
   Warranty conditions, liability, AND support -
      IF the application has been made available free OF charge, the following applies:
      * We DO NOT provide a warranty FOR Any OF the information contained in this document.
      * All other rights AND claims against Siemens AG irrespective OF legal basis are excluded. In particular claims FOR damages against Siemens AG 
      in the CASE OF Product outage, downtime, loss OF profit, either directly, indirectly OR consequential damage are excluded.
      * This does NOT apply when liability is compulsory BY law, e. g. in the CASE OF the Product liability act, premeditation, an act OF gross negligence 
      BY superiors AND managerial staff OF Siemens AG OR in cases OF fraudulent concealment OF defects.
      * This limitation OF liability also applies TO sub-contractors, suppliers, delegates, superiors AND managerial staff OF Siemens AG.
      German law shall apply TO this agreement FOR customers with head offices in Germany; Swiss law FOR customers with head offices outside Germany. 
      Application OF the United Nations Convention on Contracts FOR the International Sale OF Goods as OF 11.04.1980 (CISG) is excluded.
   *)

   // ===========================================================================
   //  Begin the LOGIC section:

   // Determine the Number of Sts_Events for given alarm/warning area
   // // S7-300 Logic:
   // UDT_Event = 66 bytes in length
   // S7-300 Logic:
   //#tempAnyPointer := #Sts_EventSummation.Sts_Events;    // temp Any Pointer for FC_ArrrayLength call.
   //"FC_ArrayLength"(ArraySource:= #tempAnyPointer, ArrayLength:=66, SIZE=> #Sts_EventSummation.Wrk_EventArraySize);
   // S7-1500 Logic:
   // "FC_ArrayLength_S7-1500"(Array_ToBe_Sized := #Sts_EventSummation.Sts_Events,
      //                      ArraySize => #Sts_EventSummation.Wrk_EventArraySize);

   // Cleanup the summation - This FB is to be called after the numerous "FB_PMLe_EventSum" calls.
   IF #Prev_NumAllEvents > #Sts_EventSummation.Sts_NumEvents THEN
       FOR #Index := #Sts_EventSummation.Sts_NumEvents TO (#Prev_NumAllEvents-1) DO
             #Sts_EventSummation.Sts_Events[#Index]:= #ZeroEvent;   // clear the first out event
       END_FOR;
   END_IF;

   #Prev_NumAllEvents := #Sts_EventSummation.Sts_NumEvents;     

   #Sts_EventSummation.Sts_Category_0_Latched := #Sts_EventSummation.Wrk_Category_0_Latched;
   #Sts_EventSummation.Sts_Category_1_Latched := #Sts_EventSummation.Wrk_Category_1_Latched;
   #Sts_EventSummation.Sts_Category_2_Latched := #Sts_EventSummation.Wrk_Category_2_Latched;
   #Sts_EventSummation.Sts_Category_3_Latched := #Sts_EventSummation.Wrk_Category_3_Latched;
   #Sts_EventSummation.Sts_Category_4_Latched := #Sts_EventSummation.Wrk_Category_4_Latched;
   #Sts_EventSummation.Sts_Category_6_Latched := #Sts_EventSummation.Wrk_Category_5_Latched;
   #Sts_EventSummation.Sts_Category_7_Latched := #Sts_EventSummation.Wrk_Category_6_Latched;
   #Sts_EventSummation.Sts_Category_8_Latched := #Sts_EventSummation.Wrk_Category_8_Latched;
   #Sts_EventSummation.Sts_Category_9_Latched := #Sts_EventSummation.Wrk_Category_9_Latched;

   #Sts_EventSummation.Sts_Category_0_NotLatched := #Sts_EventSummation.Wrk_Category_0_NotLatched;
   #Sts_EventSummation.Sts_Category_1_NotLatched := #Sts_EventSummation.Wrk_Category_1_NotLatched;
   #Sts_EventSummation.Sts_Category_2_NotLatched := #Sts_EventSummation.Wrk_Category_2_NotLatched;
   #Sts_EventSummation.Sts_Category_3_NotLatched := #Sts_EventSummation.Wrk_Category_3_NotLatched;
   #Sts_EventSummation.Sts_Category_4_NotLatched := #Sts_EventSummation.Wrk_Category_4_NotLatched;
   #Sts_EventSummation.Sts_Category_6_NotLatched := #Sts_EventSummation.Wrk_Category_5_NotLatched;
   #Sts_EventSummation.Sts_Category_7_NotLatched := #Sts_EventSummation.Wrk_Category_6_NotLatched;
   #Sts_EventSummation.Sts_Category_8_NotLatched := #Sts_EventSummation.Wrk_Category_8_NotLatched;
   #Sts_EventSummation.Sts_Category_9_NotLatched := #Sts_EventSummation.Wrk_Category_9_NotLatched;

   #Sts_EventSummation.Sts_CurrentActiveEvent  := #Sts_EventSummation.Wrk_CurrentActiveEvent; 

   //  ------------------------------------------------------------------

   ENO:= true;   // Set the ENO output
END_FUNCTION_BLOCK

FUNCTION_BLOCK "FB_TR88_CPG_EventSortFilter"   // FB3106, SCL
TITLE = PackML Event Sort Filter (TR88 CPG Template)
{ S7_Optimized_Access := 'TRUE' }
AUTHOR : FoodBev
FAMILY : ISATR88e
NAME : EvSrtFlt
VERSION : 1.21
// Sorts and filters event data. It can filter and only show events in a certain category, can sort by time, and can group by category
   VAR_INPUT
      Cmd_FilterActiveEvents : Bool;
      Cmd_FilterCategory : Bool;
      Cfg_FilterCategory : Int;
      Cmd_Sort : Bool;
      Cfg_SortCategory : Bool;
   END_VAR
   VAR_OUTPUT
      Sts_SortFilterNumEvents : Int;
   END_VAR
   VAR_IN_OUT
      In_Events : Array[0.."TR88_CPG_NoOfStsElements_EventSum"] of "UDT_TR88_CPG_Event";   // 30 Events - matches UDT declaration
      In_NumEvents : Int;
      Sts_SortFilterEventList : Array[0.."TR88_CPG_NoOfHMISortEvents"] of "UDT_TR88_CPG_Event";   // 20 Filtered Events
   END_VAR
   VAR
      Compare_True : Bool;
      temp_DT_1 : Date_And_Time;   // Temp Date & Time value #1 - Siemens
      temp_DT_2 : Date_And_Time;   // Temp Date & Time value #2 - Siemens
      FilterAcknowledged : Bool;
      FilterActive : Bool;
      FilterCategory : Bool;
      Index : Int;   // was DINT
      Index_End : Int;   // was DINT
      Index_NumEvents : Int;   // was DINT
      Index_Start : Int;   // was DINT
      MaxSize : Int;   // was DINT
      Prev_NumEvents : Int;   // was DINT
      siftDown_Child : Int;   // was DINT
      siftDown_End : Int;   // was DINT
      siftDown_Root : Int;   // was DINT
      TempEvent : "UDT_TR88_CPG_Event";
      ZeroEvent : "UDT_TR88_CPG_Event";
      Index_2 : Int;   // Index value used for DO and FOR loops
      Compare_1 : Bool;   // Siemens. Compare of TimeEvents #1
      Compare_2 : Bool;   // Siemens. Compare of TimeEvents #2
      SortingEventStatus : Array[0..29] of "UDT_TR88_CPG_Event";   // Added for V1.2
      SortingNumEventsStatus : Int;   // Added for V1.2
   END_VAR
   VAR_TEMP
      tempAnyPointer : DInt;
      siftDown_LeftChild : Int;
      siftDown_RightChild : Int;
   END_VAR
BEGIN
   // ============================================================================ 
   // FUNCTION_BLOCK "FB_PMLe_EventSortFilter"    
   // ---------------------------------------------------------------------------
   // Siemens Industry, Inc.
   // Food & Beverage VSS
   // ---------------------------------------------------------------------------
   // FUNCTIONALITY:  
   // Function Block to control Event Sort Filter commands
   // ---------------------------------------------------------------------------
   // change log table:
   // version        date          expert in charge        changes applied
   // 
   //  1.2         2012-08-20          M.Pieper             Matches Rev 1.2
   //  1.21       2015-01-27           M.Pieper            Updated S7-1500 Array Size Logic.
   // ===========================================================================
   (*
   THIS SOFTWARE IS PROVIDED "AS IS" AND WITHOUT WARRANTIES OF ANY KIND, WHETHER EXPRESS OR IMPLIED.

   General information -
       Note :  the standard applications are NOT binding AND DO NOT claim TO be complete regarding configuration, equipment OR any eventuality which may arise. 
       The standard applications DO NOT represent specific customer solutions, but are only intended TO provide support FOR typical tasks. You are responsible 
       FOR the proper operation OF the described products. These standard applications DO NOT relieve you OF your responsibility regarding the safe handling 
       when using, installing operating AND maintaining the equipment. BY using these standard applications, you agree that Siemens cannot be made liable FOR 
       possible damage beyond the mentioned liability clause. We reserve the right TO make changes AND revisions TO these standard applications at Any Time 
       without prior notice. In the CASE OF Any differences between the suggestions made in these standard applications AND other publications from Siemens, 
       such as catalogs, the contents OF the other documentation have priority.

   Warranty conditions, liability, AND support -
      IF the application has been made available free OF charge, the following applies:
      * We DO NOT provide a warranty FOR Any OF the information contained in this document.
      * All other rights AND claims against Siemens AG irrespective OF legal basis are excluded. In particular claims FOR damages against Siemens AG 
      in the CASE OF Product outage, downtime, loss OF profit, either directly, indirectly OR consequential damage are excluded.
      * This does NOT apply when liability is compulsory BY law, e. g. in the CASE OF the Product liability act, premeditation, an act OF gross negligence 
      BY superiors AND managerial staff OF Siemens AG OR in cases OF fraudulent concealment OF defects.
      * This limitation OF liability also applies TO sub-contractors, suppliers, delegates, superiors AND managerial staff OF Siemens AG.
      German law shall apply TO this agreement FOR customers with head offices in Germany; Swiss law FOR customers with head offices outside Germany. 
      Application OF the United Nations Convention on Contracts FOR the International Sale OF Goods as OF 11.04.1980 (CISG) is excluded.
   *)

   // ===========================================================================
   //  Begin the LOGIC section:
   // Event Sort and Filter
   // Determine the Number of Events for given alarm/warning area
   // UDT_Event = 66 bytes in length 
   // S7-300 Code:
   // #tempAnyPointer := #Sts_SortFilterEventList;    // temp Any Pointer for FC_ArrrayLength call.
   // "FC_ArrayLength"(ArraySource :=  #tempAnyPointer, ArrayLength := 66, SIZE =>  #MaxSize);
   // S7-1500 Code:
   "FC_ArrayLength_S7-1500"(Array_ToBe_Sized := #Sts_SortFilterEventList,
                            ArraySize => #MaxSize);

   IF #In_NumEvents < #MaxSize - 1 THEN
       #SortingNumEventsStatus := DINT_TO_INT(#In_NumEvents);
   ELSE
       #SortingNumEventsStatus := #MaxSize - 1;
   END_IF;

   // Filter
   IF #Cmd_FilterCategory OR #Cmd_FilterActiveEvents THEN
       #Index_NumEvents := 0;
       FOR #Index := 0 TO (#SortingNumEventsStatus - 1) DO         // Siemens added DINT_TO_INT   // should be "In_NumEvents-1"
           #FilterCategory := FALSE;
           #FilterAcknowledged := FALSE;
           #FilterActive := FALSE;
           IF #Cmd_FilterCategory AND (#In_Events[#Index].Category = #Cfg_FilterCategory) THEN
               #FilterCategory := 1;
           END_IF;

           IF #Cmd_FilterActiveEvents AND (#In_Events[#Index].Trigger) THEN
               #FilterActive := 1;
           END_IF;

           IF ((#Cmd_FilterCategory AND #FilterCategory) OR NOT (#Cmd_FilterCategory)) AND ((#Cmd_FilterActiveEvents AND #FilterActive) OR NOT (#Cmd_FilterActiveEvents)) THEN
               #SortingEventStatus[#Index_NumEvents] := #In_Events[#Index];
               #Index_NumEvents := #Index_NumEvents + 1;
           END_IF;

           IF (#Index_NumEvents >= #SortingNumEventsStatus) THEN
               EXIT;
           END_IF;
       END_FOR;

       #SortingNumEventsStatus := #Index_NumEvents;

       // ELSE COP(In_Events[0],Sts_SortFilterEventList[0],Sts_SortFilterNumEvents
   ELSE
       FOR #Index_2 := 0 TO #SortingNumEventsStatus - 1 DO
           #SortingEventStatus[#Index_2] := #In_Events[#Index_2];
       END_FOR;                                            // End FOR loop
   END_IF;                                                 // End Cmd_FilterCategory OR Cmd_FilterActiveEvents THEN....


   // Heap Sort #1
   IF #Cmd_Sort THEN
       // Initial Heapify
       #Index_Start := (#SortingNumEventsStatus / 2);         //-1;
       WHILE #Index_Start >= 0 DO
           // siftDown logic
           #siftDown_Root := #Index_Start;
           #siftDown_End := #SortingNumEventsStatus - 1;
           #siftDown_LeftChild := #siftDown_Root * 2 + 1;
           #siftDown_RightChild := #siftDown_Root * 2 + 2;
           WHILE (#siftDown_LeftChild) <= #siftDown_End DO //while left child exists, find which child is greatest
               IF (#siftDown_LeftChild) = #siftDown_End THEN  // if this is the last element, use it
                   #siftDown_Child := #siftDown_LeftChild;
               ELSIF #Cfg_SortCategory AND (#SortingEventStatus[#siftDown_LeftChild].Category > #SortingEventStatus[#siftDown_RightChild].Category) THEN
                   // if sorting by category, use highest category
                   #siftDown_Child := #siftDown_LeftChild;
               ELSIF (#Cfg_SortCategory AND (#SortingEventStatus[#siftDown_LeftChild].Category = #SortingEventStatus[#siftDown_RightChild].Category)) OR NOT (#Cfg_SortCategory) THEN
                   // if both children are the same cat or no sorting by cat, sort by date
                   #temp_DT_1 := #SortingEventStatus[#siftDown_LeftChild].DateTime;   // Date & Time of Event.TimeEvent[Heap]
                   #temp_DT_2 := #SortingEventStatus[#siftDown_RightChild].DateTime; // Date & Time of Event.TimeEvent[Heap+1]          
                   IF #temp_DT_1 > #temp_DT_2 THEN                                      // is [siftDown_Root*2].TimeEvent > [siftDown_Root*2+1].TimeEvent
                       #siftDown_Child := #siftDown_LeftChild;
                   ELSE
                       #siftDown_Child := #siftDown_RightChild;
                   END_IF;  // END_IF "DT1 > DT2
               ELSE
                   #siftDown_Child := #siftDown_RightChild; // this happens if right.cat > left.cat and sorting by cat
               END_IF; // END_IF "(siftDown_Root*2)..."

               //compare if root and child need to be swapped
               //swap if root has lower category or earlier date
               #Compare_True := 0;
               IF #Cfg_SortCategory AND (#SortingEventStatus[#siftDown_Root].Category < #SortingEventStatus[#siftDown_Child].Category) THEN
                   #Compare_True := 1;
               ELSIF (#Cfg_SortCategory AND (#SortingEventStatus[#siftDown_Root].Category = #SortingEventStatus[#siftDown_Child].Category))
                   OR NOT (#Cfg_SortCategory) THEN
                   #temp_DT_1 := #SortingEventStatus[#siftDown_Root].DateTime;   // Date & Time of Event.TimeEvent[Heap]
                   #temp_DT_2 := #SortingEventStatus[#siftDown_Child].DateTime;  // Date & Time of Event.TimeEvent[Heap+1] 
                   IF #temp_DT_1 < #temp_DT_2 THEN                                  // is [siftDown_Root].TimeEvent < [siftDown_Root+1].TimeEvent
                       #Compare_True := 1;
                   END_IF;  // END_IF "IF Compare_1 ..."           
               END_IF; //END_IF "IF Cfg_SortCategory AND (.."

               IF #Compare_True THEN
                   #TempEvent := #SortingEventStatus[#siftDown_Root];
                   #SortingEventStatus[#siftDown_Root] := #SortingEventStatus[#siftDown_Child];
                   #SortingEventStatus[#siftDown_Child] := #TempEvent;
                   #siftDown_Root := #siftDown_Child;
                   #siftDown_LeftChild := #siftDown_Root * 2 + 1;
                   #siftDown_RightChild := #siftDown_Root * 2 + 2;
               ELSE
                   EXIT;
               END_IF;

           END_WHILE;
           #Index_Start := #Index_Start - 1;
       END_WHILE;

       // Heap Sort #2
       #Index_End := #SortingNumEventsStatus - 1;
       WHILE #Index_End >= 1 DO
           #TempEvent := #SortingEventStatus[0];
           #SortingEventStatus[0] := #SortingEventStatus[#Index_End];
           #SortingEventStatus[#Index_End] := #TempEvent;
           // siftDown
           #siftDown_Root := 0;
           #siftDown_End := #Index_End - 1;
           #siftDown_LeftChild := #siftDown_Root * 2 + 1;
           #siftDown_RightChild := #siftDown_Root * 2 + 2;
           WHILE (#siftDown_LeftChild) <= #siftDown_End DO
               IF (#siftDown_LeftChild) = #siftDown_End THEN
                   #siftDown_Child := #siftDown_LeftChild;
               ELSIF #Cfg_SortCategory AND (#SortingEventStatus[#siftDown_LeftChild].Category > #SortingEventStatus[#siftDown_RightChild].Category) THEN
                   #siftDown_Child := #siftDown_LeftChild;
               ELSIF (#Cfg_SortCategory AND (#SortingEventStatus[#siftDown_LeftChild].Category = #SortingEventStatus[#siftDown_RightChild].Category)) OR NOT (#Cfg_SortCategory) THEN
                   #temp_DT_1 := #SortingEventStatus[#siftDown_LeftChild].DateTime;
                   #temp_DT_2 := #SortingEventStatus[#siftDown_RightChild].DateTime;

                   IF #temp_DT_1 > #temp_DT_2 THEN
                       #siftDown_Child := #siftDown_LeftChild;
                   ELSE
                       #siftDown_Child := #siftDown_RightChild;
                   END_IF;
               ELSE
                   #siftDown_Child := #siftDown_RightChild;
               END_IF;

               #Compare_True := FALSE;
               IF #Cfg_SortCategory AND (#SortingEventStatus[#siftDown_Root].Category < #SortingEventStatus[#siftDown_Child].Category) THEN
                   #Compare_True := TRUE;
               ELSIF (#Cfg_SortCategory AND (#SortingEventStatus[#siftDown_Root].Category = #SortingEventStatus[#siftDown_Child].Category)) OR NOT (#Cfg_SortCategory) THEN
                   #temp_DT_1 := #SortingEventStatus[#siftDown_Root].DateTime;
                   #temp_DT_2 := #SortingEventStatus[#siftDown_Child].DateTime;

                   IF #temp_DT_1 < #temp_DT_2 THEN
                       #Compare_True := TRUE;
                   END_IF;
               END_IF;

               IF #Compare_True THEN
                   #TempEvent := #SortingEventStatus[#siftDown_Root];
                   #SortingEventStatus[#siftDown_Root] := #SortingEventStatus[#siftDown_Child];
                   #SortingEventStatus[#siftDown_Child] := #TempEvent;
                   #siftDown_Root := #siftDown_Child;
                   #siftDown_LeftChild := #siftDown_Root * 2 + 1;
                   #siftDown_RightChild := #siftDown_Root * 2 + 2;
               ELSE
                   EXIT;
               END_IF;
           END_WHILE;
           #Index_End := #Index_End - 1;
       END_WHILE;
   END_IF; //END_IF -> IF Cmd_Sort THEN"

   // Copy SortingEventStatus (working area) to Sts_SortFilterEventList (out)
   // FOR Index  := 0  TO SortingNumEventsStatus DO   
   FOR #Index := 0 TO #SortingNumEventsStatus - 1 DO
       #Sts_SortFilterEventList[#Index] := #SortingEventStatus[#Index];
   END_FOR;
   // End FOR loop
   #Sts_SortFilterNumEvents := #SortingNumEventsStatus;

   // Clean up event list
   IF #Prev_NumEvents > #Sts_SortFilterNumEvents THEN
       //FOR Index  :=  Sts_SortFilterNumEvents TO Prev_NumEvents-1 DO
       FOR #Index := #Sts_SortFilterNumEvents TO #Prev_NumEvents DO
           #Sts_SortFilterEventList[#Index] := #ZeroEvent;
       END_FOR;
   END_IF;

   #Prev_NumEvents := #Sts_SortFilterNumEvents;

   // End of Main Logic.
   //----------------------------------------------------- 

   ENO := true;   // Set the ENO output
END_FUNCTION_BLOCK

FUNCTION_BLOCK "FB_TR88_CPG_Msg_Scroll"   // FB3108, SCL
TITLE = PackML HMI Message Scroll (TR88 CPG Template)
{ S7_Optimized_Access := 'TRUE' }
AUTHOR : FoodBev
FAMILY : ISATR88e
NAME : MsgScrll
VERSION : 1.0
   VAR_INPUT
      Trigger : Bool;   // input trigger to enable scroll logic
      NumEvents : Int;   // input value with number of active events
      In_Events : Array[0.."TR88_CPG_NoOfHMISortEvents"] of "UDT_TR88_CPG_Event";   // incoming events list
   END_VAR
   VAR_OUTPUT
      Msg_Scroll : String[40];   // message output value
   END_VAR
   VAR
      Scroll_Index : Int;   // index value for scroll logic
      TriggerOS : Bool;
      MaxSize : Int;   // was DINT
   END_VAR
   VAR_TEMP
      Scroll_Index_Max : Int;
   END_VAR
BEGIN
   // ============================================================================ 
   // FUNCTION_BLOCK "FB_PMLe_Msg_Scroll"    
   // ---------------------------------------------------------------------------
   // Siemens Industry, Inc.
   // Food & Beverage VMM
   // ---------------------------------------------------------------------------
   // functionality:
   // Function Block used to scoll messages from an array of EVENT to a single
   // ---------------------------------------------------------------------------
   // change log table:
   // version        date          expert in charge        changes applied
   // 
   // 1.0         2012-02-28          M.Pieper           Matches Rev 1.0
   // 1.01        2015-04-01          M.Pieper          Changed "In_Events" from array size of [0..19]
   //                                                    to Array[0.."CPG_TR88_NoOfHMISortEvents"]
   // ===========================================================================
   (*
   THIS SOFTWARE IS PROVIDED "AS IS" AND WITHOUT WARRANTIES OF ANY KIND, WHETHER EXPRESS OR IMPLIED.

   General information -
       Note :  the standard applications are NOT binding AND DO NOT claim TO be complete regarding configuration, equipment OR any eventuality which may arise. 
       The standard applications DO NOT represent specific customer solutions, but are only intended TO provide support FOR typical tasks. You are responsible 
       FOR the proper operation OF the described products. These standard applications DO NOT relieve you OF your responsibility regarding the safe handling 
       when using, installing operating AND maintaining the equipment. BY using these standard applications, you agree that Siemens cannot be made liable FOR 
       possible damage beyond the mentioned liability clause. We reserve the right TO make changes AND revisions TO these standard applications at Any Time 
       without prior notice. In the CASE OF Any differences between the suggestions made in these standard applications AND other publications from Siemens, 
       such as catalogs, the contents OF the other documentation have priority.

   Warranty conditions, liability, AND support -
      IF the application has been made available free OF charge, the following applies:
      * We DO NOT provide a warranty FOR Any OF the information contained in this document.
      * All other rights AND claims against Siemens AG irrespective OF legal basis are excluded. In particular claims FOR damages against Siemens AG 
      in the CASE OF Product outage, downtime, loss OF profit, either directly, indirectly OR consequential damage are excluded.
      * This does NOT apply when liability is compulsory BY law, e. g. in the CASE OF the Product liability act, premeditation, an act OF gross negligence 
      BY superiors AND managerial staff OF Siemens AG OR in cases OF fraudulent concealment OF defects.
      * This limitation OF liability also applies TO sub-contractors, suppliers, delegates, superiors AND managerial staff OF Siemens AG.
      German law shall apply TO this agreement FOR customers with head offices in Germany; Swiss law FOR customers with head offices outside Germany. 
      Application OF the United Nations Convention on Contracts FOR the International Sale OF Goods as OF 11.04.1980 (CISG) is excluded.
   *)

   // ===========================================================================
   //  Begin the LOGIC section:
   "FC_ArrayLength_S7-1500"(Array_ToBe_Sized := #In_Events,
                            ArraySize => #MaxSize);

   IF #NumEvents > #MaxSize THEN
       #Scroll_Index_Max := #MaxSize;
   ELSE
       #Scroll_Index_Max := #NumEvents;
   END_IF;

   // Statement Section 
   IF #Trigger AND NOT #TriggerOS THEN
       #Scroll_Index := #Scroll_Index + 1;  // increment the indext
       IF  #Scroll_Index > #Scroll_Index_Max - 1 THEN
               #Scroll_Index := 0;
           END_IF;
      #Msg_Scroll := #In_Events[#Scroll_Index].Message;      // move the message from the UDT_Event structure to string output.  

       #TriggerOS := TRUE;              // Set the trigger OS bit
   END_IF;

   IF NOT #Trigger AND #TriggerOS THEN
       #TriggerOS := FALSE;
   END_IF;

   ENO:= true;   // Set the ENO output
END_FUNCTION_BLOCK

FUNCTION_BLOCK "FB_TR88_CPG_OEE"   // FB3109, SCL
TITLE = PackML Real-Time OEE Calculation (TR88 CPG Template)
{ S7_Optimized_Access := 'TRUE' }
AUTHOR : FoodBev
FAMILY : ISATR88
NAME : OEE
VERSION : 1.1
   VAR_INPUT
      TotalProdProcessed : DInt;   // Total Number OF Products Processed
      TotalDefectiveProd : DInt;   // Total Number OF Defective Products
      TimeSinceLastReset : DInt;   // Total Acumulative TIME since Last RESET
      MachineDesignSpeed : Real;   // Machine Design Speed
   END_VAR
   VAR_OUTPUT
      OEE_RealTimeValue : Real;   // REAL TIME OEE value (availabilty x performance x quality)
      OEE_Availability : Real;   // OEE - Availability value
      OEE_Performance : Real;   // OEE - Performance value
      OEE_Quality : Real;   // OEE - Quality value
   END_VAR
   VAR_IN_OUT
      ModeCumulativeTimes : Array[0.."LPMLV30_MODES_UPPER_LIM"] of DInt;   // Mode Cummulative Times
   END_VAR
   VAR
      TotalProdProcessed_In : DInt;   // Initial "TotalProdProcessed" value after accum TIME reset
      TotalDefectiveProd_In : DInt;   // Initial "TotalDefectiveProcessed" value after accum TIME reset
      AcumTimeEqualZero : Bool;   // The "TimeSinceLastReset" is = 0 seconds
      AcumTimeEqualZeroOS : Bool;   // OneShot for "TimeSinceLastReset" is = 0 seconds
   END_VAR
   VAR_TEMP
      temp_TimeSinceLastReset : Real;   // used to eliminate divide by zero errors
      temp_TotalProducts : Real;   // used to eliminate divide by zero errors
      temp_DefectiveProducts : Real;   // used to eliminate divide by zero errors
   END_VAR
BEGIN
   // ============================================================================ 
   // FUNCTION_BLOCK "FB_PML_OEE"    
   // ---------------------------------------------------------------------------
   // Siemens Industry, Inc.
   // Food & Beverage VSS
   // ---------------------------------------------------------------------------
   // functionality: Function Block to calculate real-time OEE values
   // ---------------------------------------------------------------------------
   // change log table:
   // version        date          expert in charge        changes applied
   // 
   //  1.00         2012-02-28          M.Pieper        Original - using OEE Realtime calculation
   //  1.10         2012-09-04          M.Pieper        Added seperate Availabity, Performace, Quality calculation
   //  1.20         2014-07-07          M.Pieper        Updated interface FOR new Mode/State FB          
   //  1.201        2016-03-01          M.Pieper        Added logic to prevent floating point / divide by zero errors
   //  // ===========================================================================
   (*
   THIS SOFTWARE IS PROVIDED "AS IS" AND WITHOUT WARRANTIES OF ANY KIND, WHETHER EXPRESS OR IMPLIED.

   General information -
       Note :  the standard applications are NOT binding AND DO NOT claim TO be complete regarding configuration, equipment OR any eventuality which may arise. 
       The standard applications DO NOT represent specific customer solutions, but are only intended TO provide support FOR typical tasks. You are responsible 
       FOR the proper operation OF the described products. These standard applications DO NOT relieve you OF your responsibility regarding the safe handling 
       when using, installing operating AND maintaining the equipment. BY using these standard applications, you agree that Siemens cannot be made liable FOR 
       possible damage beyond the mentioned liability clause. We reserve the right TO make changes AND revisions TO these standard applications at Any Time 
       without prior notice. In the CASE OF Any differences between the suggestions made in these standard applications AND other publications from Siemens, 
       such as catalogs, the contents OF the other documentation have priority.

   Warranty conditions, liability, AND support -
      IF the application has been made available free OF charge, the following applies:
      * We DO NOT provide a warranty FOR Any OF the information contained in this document.
      * All other rights AND claims against Siemens AG irrespective OF legal basis are excluded. In particular claims FOR damages against Siemens AG 
      in the CASE OF Product outage, downtime, loss OF profit, either directly, indirectly OR consequential damage are excluded.
      * This does NOT apply when liability is compulsory BY law, e. g. in the CASE OF the Product liability act, premeditation, an act OF gross negligence 
      BY superiors AND managerial staff OF Siemens AG OR in cases OF fraudulent concealment OF defects.
      * This limitation OF liability also applies TO sub-contractors, suppliers, delegates, superiors AND managerial staff OF Siemens AG.
      German law shall apply TO this agreement FOR customers with head offices in Germany; Swiss law FOR customers with head offices outside Germany. 
      Application OF the United Nations Convention on Contracts FOR the International Sale OF Goods as OF 11.04.1980 (CISG) is excluded.
   *)

   // ===========================================================================
   //  Begin the LOGIC section:
   //  
   (* ISA TR88.00.02 Document - 9.1 OEE Definition:
   Overall Equipment Effectiveness (OEE) is a measure comparing how well manufacturing equipment is running compared to the ideal plant. The resulting measurement is expressed as the ratio of the actual
   output of the equipment divided by the maximum possible output of the equipment under ideal conditions. OEE is calculated by multiplying three independently measured values: Availability,
   Performance Rate, and Quality Rate. The fundamental OEE definition is defined as an availability ratio multiplied by a performance ratio multiplied by a quality ratio.

   OEE = Availability x Performance x Quality

   Where each component is defined as the following:
   Availability = Operating Time / Planned Production Time
   Performance = Total Pieces / (Operating Time* Ideal Run Rate)
   Quality = Good Pieces / Total Pieces

   OEE is often displayed as a waterfall object in which the major components of Availability, Performance, and Quality are displayed graphically.
   *)

   // Determine is TimeSinceLastReset value is equal to zero.
   IF  #TimeSinceLastReset   = 0 THEN
       #AcumTimeEqualZero   := TRUE;  // SET the AcumTimeEqualZero bool tag
   ELSE
       #AcumTimeEqualZero   := FALSE; // RESET the AcumTimeEqualZero bool tag
       #AcumTimeEqualZeroOS := FALSE; // RESET the AcumTimeEqualZero one-shot bool tag
   END_IF;

   // Update the AcumTimeEqualZeroOS One-Shot bool
   IF #AcumTimeEqualZero AND NOT #AcumTimeEqualZeroOS THEN
      #AcumTimeEqualZeroOS := TRUE;  // Set the One-Shot bool tag
   END_IF;

   // Update the inital product count values after the accum timer value has been reset
   IF #AcumTimeEqualZeroOS THEN
      #TotalProdProcessed_In := #TotalProdProcessed;
      #TotalDefectiveProd_In := #TotalDefectiveProd;
   END_IF;  

   // Update the TimeSinceLastReset temp. value.  If = 0 (zero) then change to 0.0001 to ensure no divide by zero errors
   IF #TimeSinceLastReset = 0 THEN
       #temp_TimeSinceLastReset := 0.0001;
   ELSE
       #temp_TimeSinceLastReset := DINT_TO_REAL(#TimeSinceLastReset);
   END_IF;

   (*  9.1.1 Availability Definition
   Availability is defined as operating time divided by planned production time. The basic concept behind availability is to show the time the machine has been running divided by the time that the
   machine has been planned to run. Typical losses in this area are losses to unplanned maintenance, cleaning, changeovers, and breakdowns.
   * Availability = Operating Time / Planned Production Time Operating Time is defined as the amount of time the machine has been attempting to produce parts.  
   * Planned Production Time is defined as the total amount of time the machine has been scheduled to run. 
   *)
   // Availablity = operating time (attempt to run production) / planned production time
   #OEE_Availability :=   DINT_TO_REAL (#ModeCumulativeTimes[1]) / #temp_TimeSinceLastReset;
   IF #OEE_Availability > 1 THEN #OEE_Availability := 1.0; END_IF;
   IF #OEE_Availability < 0 THEN #OEE_Availability := 0.0; END_IF;

   (* 9.1.2 Performance Definition
   Performance is defined as the total number of pieces on which the machine operated divided by the ideal production if a machine ran perfectly for the allocated amount of operating time.
   * Performance = Total Pieces / (Operating Time* Ideal Run Rate).  
   * Total Pieces is defined as good pieces and bad pieces during the production run. This should be linked to the main consumed count of the machine. If a filler, this should be bottles into the filler.
   * Operating Time is defined as the amount of time the machine has been attempting to produce parts. (Same as above)
   * Ideal Run Rate is defined as the ideal rate that the machine can run for the product that is being run on the machine and the way the machine is configured.
   *)
   // Performance = Total Pieces / (Operating Time * Ideal Run Rate / 60)
   #OEE_Performance := (DINT_TO_REAL(#TotalProdProcessed-#TotalProdProcessed_In))/((#temp_TimeSinceLastReset * #MachineDesignSpeed/60.0));
   IF #OEE_Performance > 1 THEN #OEE_Performance := 1.0; END_IF;
   IF #OEE_Performance < 0 THEN #OEE_Performance := 0.0; END_IF;

   (*  9.1.3 Quality Definition
   Quality is defined as the total number of good pieces divided by the total number of pieces on which the machine operated.
   * Quality = Good Pieces / Total Pieces
   * Good Pieces is defined as only good pieces processed during the production run. So this is the main production processed count of the machine. If a filler, this should be bottles out of the filler.
   * Total Pieces includes good pieces and bad pieces during the production run. This should be linked to the main consumed count of the machine. 
      If a filler, this should be bottles into the filler. This should be the same count as used in the performance definition.
   *)
   // Quality = Good Piece / Total Piece
   #temp_TotalProducts     :=  DINT_TO_REAL(#TotalProdProcessed-#TotalProdProcessed_In);
   #temp_DefectiveProducts :=  DINT_TO_REAL(#TotalDefectiveProd-#TotalDefectiveProd_In);

   // Prevent divide by zero errors by checking if Total Products <> 0.0
   IF (#TotalProdProcessed-#TotalProdProcessed_In) = 0 THEN 
       #temp_TotalProducts := 0.0001;
   END_IF;

   // Make sure that defective products < total products
   IF #temp_DefectiveProducts > #temp_TotalProducts THEN
       #temp_DefectiveProducts := 0.0;
   END_IF;

   #OEE_Quality            := (#temp_TotalProducts - #temp_DefectiveProducts) / #temp_TotalProducts;
   IF #OEE_Quality  > 1 THEN #OEE_Quality  := 1.0; END_IF;
   IF #OEE_Quality  < 0 THEN #OEE_Quality  := 0.0; END_IF;
   IF #temp_TotalProducts  = 0 THEN #OEE_Quality  := 0.0; END_IF;

   // OEE_ReatTimeValue := ((DINT_TO_REAL(TotalProdProcessed-TotalProdProcessed_Initial) - DINT_TO_REAL(TotalDefectiveProd-TotalDefectiveProd_Initial)) / ((DINT_TO_REAL(TimeSinceLastReset) * MachineDesignSpeed/60.0)));
   #OEE_RealTimeValue := #OEE_Availability * #OEE_Performance * #OEE_Quality;

   // End of Main Logic.
   ENO:= true;   // Set the ENO output
END_FUNCTION_BLOCK

FUNCTION_BLOCK "FB_TR88_CPG_AlarmMove"   // FB3110, SCL
TITLE = PackML Alarm Move
{ S7_Optimized_Access := 'TRUE' }
AUTHOR : FoodBev
FAMILY : ISATR88e
NAME : AlrmMov
VERSION : 1.01
// ------------------------------------------------------------------------------------------
//   Begin the variable declartion section ....
//  Block Parameters
   VAR_INPUT
      Sts_NumEvents : Int;   // Number OF Active Alarms
   END_VAR
   VAR_OUTPUT
      Sts_error : Bool;   // Error Status. 0=no error, 1=error
      Sts_errorCode : Int;   // Error code /number
   END_VAR
   VAR_IN_OUT
      Source : Array[0.."TR88_CPG_NoOfStsElements_EventSum"] of "UDT_TR88_CPG_Event";   // source location of the machine alarms
      Destination : Array[0.."TR88_CPG_NoOfPackTagsAdminEvents"] of "UDT_TR88_CPG_Event";   // destination location of the PackTag alarms
   END_VAR
   VAR
      Source_NumEvents : Int;   // MAX # OF Events - source event list
      Destination_NumEvents : Int;   // MAX # OF Events - destination event list
      Index : Int;   // index value
      Prev_NumEvents : Int;   // previous number OF events
      ZeroEvent : "UDT_TR88_CPG_Event";   // blank event
      Wrk_NumEvents : Int;   // working number of active events
   END_VAR
   VAR_TEMP
      tempAnyPointer : DInt;
   END_VAR
BEGIN
   // ============================================================================ 
   // FUNCTION_BLOCK "FB_AlarmMove"    
   // ---------------------------------------------------------------------------
   // Siemens Industry, Inc.
   // Food & Beverage VSS
   // ---------------------------------------------------------------------------
   // functionality:
   // Function Block to move alrm structures
   // ---------------------------------------------------------------------------
   // change log table:
   // version        date          expert in charge        changes applied
   // 
   //  1.00         2012-02-28          M.Pieper        Original -
   //  1.01         2015-01-27          M.Pieper        Added S7-1500 logic to determine array sizes
   // ===========================================================================
   (*
   THIS SOFTWARE IS PROVIDED "AS IS" AND WITHOUT WARRANTIES OF ANY KIND, WHETHER EXPRESS OR IMPLIED.

   General information -
       Note :  the standard applications are NOT binding AND DO NOT claim TO be complete regarding configuration, equipment OR any eventuality which may arise. 
       The standard applications DO NOT represent specific customer solutions, but are only intended TO provide support FOR typical tasks. You are responsible 
       FOR the proper operation OF the described products. These standard applications DO NOT relieve you OF your responsibility regarding the safe handling 
       when using, installing operating AND maintaining the equipment. BY using these standard applications, you agree that Siemens cannot be made liable FOR 
       possible damage beyond the mentioned liability clause. We reserve the right TO make changes AND revisions TO these standard applications at Any Time 
       without prior notice. In the CASE OF Any differences between the suggestions made in these standard applications AND other publications from Siemens, 
       such as catalogs, the contents OF the other documentation have priority.

   Warranty conditions, liability, AND support -
      IF the application has been made available free OF charge, the following applies:
      * We DO NOT provide a warranty FOR Any OF the information contained in this document.
      * All other rights AND claims against Siemens AG irrespective OF legal basis are excluded. In particular claims FOR damages against Siemens AG 
      in the CASE OF Product outage, downtime, loss OF profit, either directly, indirectly OR consequential damage are excluded.
      * This does NOT apply when liability is compulsory BY law, e. g. in the CASE OF the Product liability act, premeditation, an act OF gross negligence 
      BY superiors AND managerial staff OF Siemens AG OR in cases OF fraudulent concealment OF defects.
      * This limitation OF liability also applies TO sub-contractors, suppliers, delegates, superiors AND managerial staff OF Siemens AG.
      German law shall apply TO this agreement FOR customers with head offices in Germany; Swiss law FOR customers with head offices outside Germany. 
      Application OF the United Nations Convention on Contracts FOR the International Sale OF Goods as OF 11.04.1980 (CISG) is excluded.
   *)

   // ===========================================================================
   //  Begin the LOGIC section:

   // Determine the Number of Sts_Events for given alarm/warning are
   // UDT_Event = 66 bytes in length
   // S7-300 Code:
   //#tempAnyPointer := #Source;    // temp Any Pointer for FC_ArrrayLength call.
   //"FC_ArrayLength"(ArraySource:= #tempAnyPointer, ArrayLength:=66, SIZE=> #Source_NumEvents);
   //
   //#tempAnyPointer := #Destination;    // temp Any Pointer for FC_ArrrayLength call.
   //"FC_ArrayLength"(ArraySource:= #tempAnyPointer, ArrayLength:=66, SIZE=> #Destination_NumEvents);
   //
   // S7-1500 Code:
   "FC_ArrayLength_S7-1500"(Array_ToBe_Sized := #Source,
                            ArraySize => #Source_NumEvents);

   "FC_ArrayLength_S7-1500"(Array_ToBe_Sized := #Destination,
                            ArraySize => #Destination_NumEvents);

   #Wrk_NumEvents := #Sts_NumEvents;

   IF (#Destination_NumEvents < #Source_NumEvents) AND (#Destination_NumEvents < #Sts_NumEvents) THEN
       #Wrk_NumEvents :=#Destination_NumEvents;
   END_IF;

   IF (#Source_NumEvents < #Destination_NumEvents) AND (#Source_NumEvents < #Sts_NumEvents) THEN
      #Wrk_NumEvents :=#Source_NumEvents;
   END_IF;


   FOR #Index  := 0  TO #Wrk_NumEvents - 1 DO           
     #Destination[#Index]  := #Source[#Index];
   END_FOR;

   // Clean up event list

   IF #Prev_NumEvents > #Wrk_NumEvents  THEN
       //FOR Index  :=  Sts_SortFilterNumEvents TO Prev_NumEvents-1 DO
       FOR #Index  :=  #Wrk_NumEvents TO #Prev_NumEvents DO
           #Destination[#Index+1]  :=  #ZeroEvent;
       END_FOR;
   END_IF;

   #Prev_NumEvents := #Wrk_NumEvents; 


   //  ------------------------------------------------------------------

   ENO:= true;   // Set the ENO output
END_FUNCTION_BLOCK

FUNCTION_BLOCK "FB_TR88_CPG_AlarmHistory"   // FB3111, SCL
TITLE = PackML Alarm History (TR88 CPG Template)
{ S7_Optimized_Access := 'TRUE' }
AUTHOR : FoodBev
FAMILY : ISATR88
NAME : AlrmHist
VERSION : 1.0
   VAR_IN_OUT
      In_StopReasonAlarm : "UDT_TR88_CPG_Event";   // Input - Stop Reason Alarm (structure)
      Sts_AlarmHistory : Array[0.."TR88_CPG_NoOfPackTagsAdminEventHistory"] of "UDT_TR88_CPG_Event";   // Status- Alarm History Log
   END_VAR
   VAR
      AlarmArraySize : Int;   // Max # of Events in the Alarm History Array
      TriggerOS_Pos : Bool;   // Trigger One Shot - positve edge
      TriggerOS_Neg : Bool;   // Trigger One Shot - negative edge
      error_RTC : Int;   // Error code for reading of Real Time Clock
      Event_CurDateTime : Date_And_Time;   // temp value for current date & time
      FB_1stScanBit : Bool;   // 0=1st scan of FB; set to 1 after 1st FB scan...
   END_VAR
   VAR_TEMP
      Index : Int;
   END_VAR
   VAR CONSTANT
      Zero : Int := 0;
      NegativeOne : Int := -1;
   END_VAR
BEGIN
   // ============================================================================ 
   // FUNCTION_BLOCK "FB_PML_AlarmHistory"
   // ---------------------------------------------------------------------------
   // Siemens Industry, Inc.
   // Food & Beverage VSS
   // ---------------------------------------------------------------------------
   // FUNCTIONALITY:  
   // FUNCTION Block used to capture the current Stop ReasonAlarm (i.e. 'Machine
   //    First Fault') to the PackTags AlarmHistory log.
   // 
   // ---------------------------------------------------------------------------
   // change log table:
   // version        date          expert in charge        changes applied
   //  1.0       2014-12-15         Mike Pieper            
   //  
   //  ===========================================================================
   (*
   THIS SOFTWARE IS PROVIDED "AS IS" AND WITHOUT WARRANTIES OF ANY KIND, WHETHER EXPRESS OR IMPLIED.

   General information -
       Note :  the standard applications are NOT binding AND DO NOT claim TO be complete regarding configuration, equipment OR any eventuality which may arise. 
       The standard applications DO NOT represent specific customer solutions, but are only intended TO provide support FOR typical tasks. You are responsible 
       FOR the proper operation OF the described products. These standard applications DO NOT relieve you OF your responsibility regarding the safe handling 
       when using, installing operating AND maintaining the equipment. BY using these standard applications, you agree that Siemens cannot be made liable FOR 
       possible damage beyond the mentioned liability clause. We reserve the right TO make changes AND revisions TO these standard applications at Any Time 
       without prior notice. In the CASE OF Any differences between the suggestions made in these standard applications AND other publications from Siemens, 
       such as catalogs, the contents OF the other documentation have priority.

   Warranty conditions, liability, AND support -
      IF the application has been made available free OF charge, the following applies:
      * We DO NOT provide a warranty FOR Any OF the information contained in this document.
      * All other rights AND claims against Siemens AG irrespective OF legal basis are excluded. In particular claims FOR damages against Siemens AG 
      in the CASE OF Product outage, downtime, loss OF profit, either directly, indirectly OR consequential damage are excluded.
      * This does NOT apply when liability is compulsory BY law, e. g. in the CASE OF the Product liability act, premeditation, an act OF gross negligence 
      BY superiors AND managerial staff OF Siemens AG OR in cases OF fraudulent concealment OF defects.
      * This limitation OF liability also applies TO sub-contractors, suppliers, delegates, superiors AND managerial staff OF Siemens AG.
      German law shall apply TO this agreement FOR customers with head offices in Germany; Swiss law FOR customers with head offices outside Germany. 
      Application OF the United Nations Convention on Contracts FOR the International Sale OF Goods as OF 11.04.1980 (CISG) is excluded.
   *)

   // ===========================================================================
   //  Begin the LOGIC section:
   // 
   // Frist Scan Logic
   IF #FB_1stScanBit = 0 THEN
       "FC_ArrayLength_S7-1500"(Array_ToBe_Sized := #Sts_AlarmHistory,
                                ArraySize => #AlarmArraySize);
       #FB_1stScanBit:=1;      // Set the FB 1st Scan Bit
   END_IF;

   // Positive Trigger
   IF #In_StopReasonAlarm.Trigger = 1 AND #TriggerOS_Pos = 0 THEN
       // execute code for new incoming event
       #TriggerOS_Pos:= 1;                 // Set the OS bit 

       // Index the existing Alarm History Array (FIFO).
       FOR #Index := #AlarmArraySize-1 TO 1 BY -1 DO
           #Sts_AlarmHistory[#Index] := #Sts_AlarmHistory[#Index-1];
       END_FOR;

       // Update the Array[0] with the current alarm information
       #Sts_AlarmHistory[0] := #In_StopReasonAlarm;

       END_IF;

       IF #In_StopReasonAlarm.Trigger = FALSE AND #TriggerOS_Pos = TRUE THEN
           // Reset the OS Bit
           #TriggerOS_Pos := FALSE;                 // Reset the OS bit   
       END_IF;

       // Negative Trigger
       IF #In_StopReasonAlarm.Trigger = 0 AND #TriggerOS_Neg = 0 THEN
           // execute code for new incoming event
           #TriggerOS_Neg := TRUE;                 // Set the OS bit 
           // Capture the Alarm Ack. Time.
           #error_RTC := RD_SYS_T(OUT => #Event_CurDateTime);            // Read the Real Time Clock
               #error_RTC := RD_SYS_T(OUT => #Event_CurDateTime);            // Read the Real Time Clock
           #Sts_AlarmHistory[0].AckDateTime := #Event_CurDateTime; // update Acknowledge time.TimeAck := #Event_CurDateTime; // update Acknowledge time

       END_IF;

       IF #In_StopReasonAlarm.Trigger = 1 AND #TriggerOS_Pos = 1 THEN
           // Reset the OS Bit
           #TriggerOS_Neg := 0;                 // Reset the OS bit   
       END_IF;

       //----------------------------------------------------- 
       ENO := true;   // Set the ENO output
END_FUNCTION_BLOCK

FUNCTION "FC_ArrayLength_S7-1500" : Void   // FC3102, SCL
TITLE = FC used to determine the length of an array (as a FC call)
{ S7_Optimized_Access := 'TRUE' }
AUTHOR : FoodBev
FAMILY : ISATR88
NAME : AryLen
VERSION : 1.1
// Changed to "#ArraySize :=
   VAR_INPUT
      Array_ToBe_Sized : Variant;   // Array to be sized
   END_VAR
   VAR_OUTPUT
      ArraySize : Int;   // Number of elements (size) in an array
   END_VAR
   VAR_TEMP
      temp_UDint : UDInt;
   END_VAR
BEGIN
   // ============================================================================ 
   // FUNCTION_BLOCK "FC_ArrayLength_S7-1500"    
   // ---------------------------------------------------------------------------
   // Siemens Industry, Inc.
   // Food & Beverage VSS
   // ---------------------------------------------------------------------------
   // Functionality:
   // Function Call to determine the length of any array
   //  using optimized S7-1x00 Data Blocks (DB)  
   // ---------------------------------------------------------------------------
   // change log table:
   // version        date          expert in charge        changes applied
   // 
   //  1.00         2014-12-08         M.Pieper            Inital Release - 
   // ===========================================================================
   (*
   THIS SOFTWARE IS PROVIDED "AS IS" AND WITHOUT WARRANTIES OF ANY KIND, WHETHER EXPRESS OR IMPLIED.

   General information -
       Note :  the standard applications are NOT binding AND DO NOT claim TO be complete regarding configuration, equipment OR any eventuality which may arise. 
       The standard applications DO NOT represent specific customer solutions, but are only intended TO provide support FOR typical tasks. You are responsible 
       FOR the proper operation OF the described products. These standard applications DO NOT relieve you OF your responsibility regarding the safe handling 
       when using, installing operating AND maintaining the equipment. BY using these standard applications, you agree that Siemens cannot be made liable FOR 
       possible damage beyond the mentioned liability clause. We reserve the right TO make changes AND revisions TO these standard applications at Any Time 
       without prior notice. In the CASE OF Any differences between the suggestions made in these standard applications AND other publications from Siemens, 
       such as catalogs, the contents OF the other documentation have priority.

